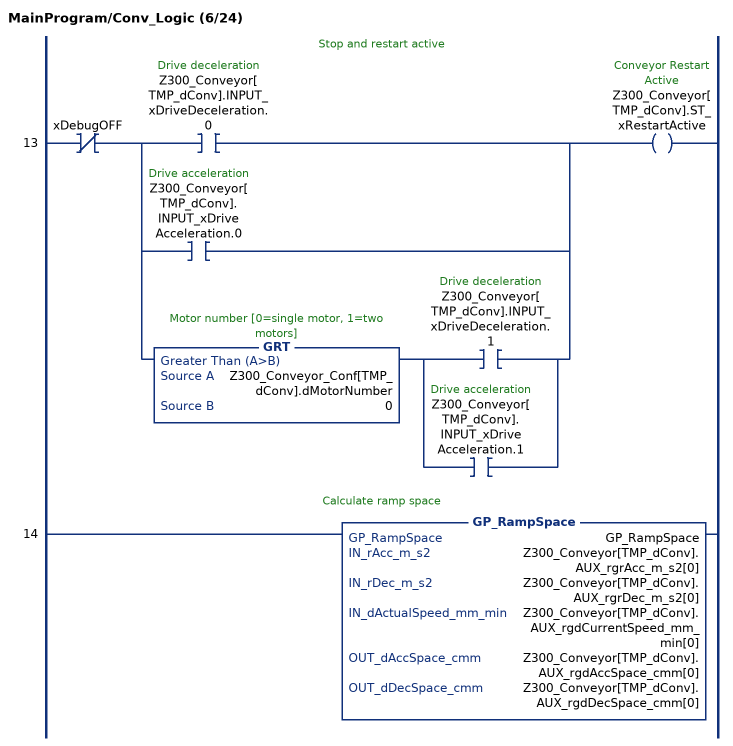
   // Stop and restart active
   13: XIO(xDebugOFF)[[XIC(Z300_Conveyor[TMP_dConv].INPUT_xDriveDeceleration.0) ,XIC(Z300_Conveyor[TMP_dConv].INPUT_xDriveAcceleration.0) ] ,GRT(Z300_Conveyor_Conf[TMP_dConv].dMotorNumber,0) [XIC(Z300_Conveyor[TMP_dConv].INPUT_xDriveDeceleration.1) ,XIC(Z300_Conveyor[TMP_dConv].INPUT_xDriveAcceleration.1) ] ]OTE(Z300_Conveyor[TMP_dConv].ST_xRestartActive);
   // Calculate ramp space
   14: GP_RampSpace(GP_RampSpace,Z300_Conveyor[TMP_dConv].AUX_rgrAcc_m_s2[0],Z300_Conveyor[TMP_dConv].AUX_rgrDec_m_s2[0],Z300_Conveyor[TMP_dConv].AUX_rgdCurrentSpeed_mm_min[0],Z300_Conveyor[TMP_dConv].AUX_rgdAccSpace_cmm[0],Z300_Conveyor[TMP_dConv].AUX_rgdDecSpace_cmm[0]);
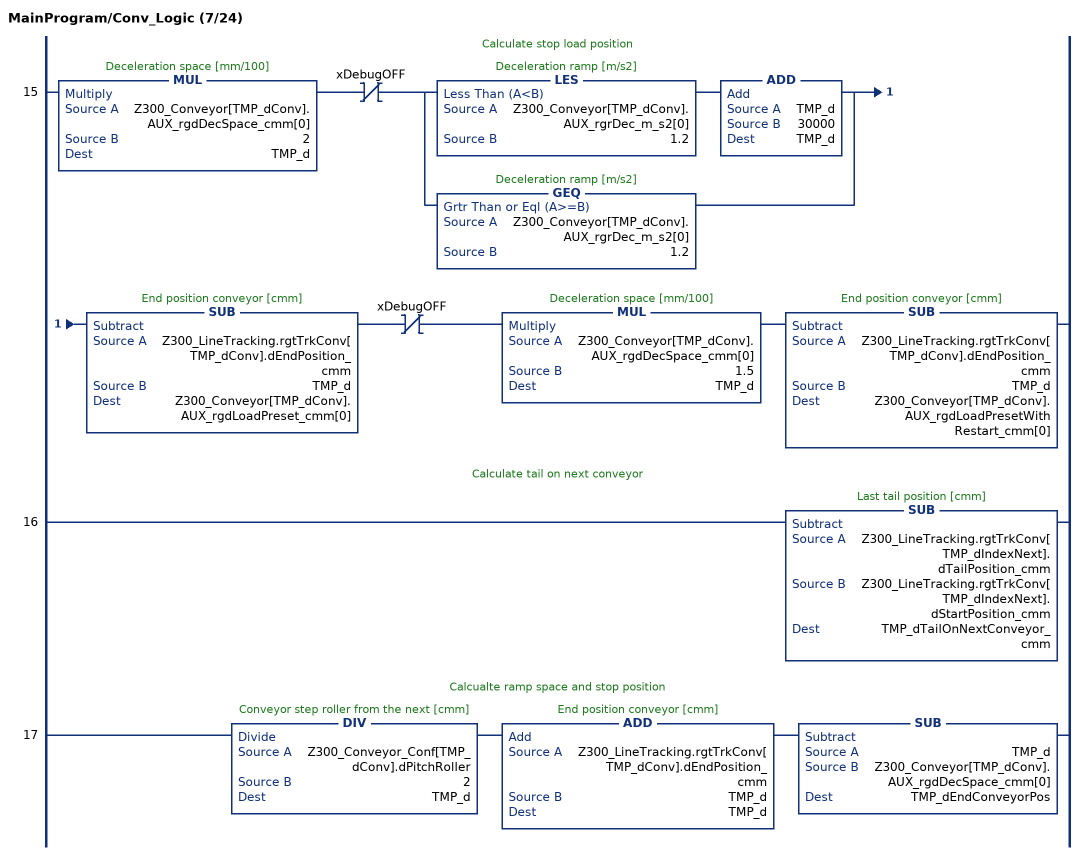
   // Calculate stop load position
   15: MUL(Z300_Conveyor[TMP_dConv].AUX_rgdDecSpace_cmm[0],2,TMP_d)XIO(xDebugOFF)[LES(Z300_Conveyor[TMP_dConv].AUX_rgrDec_m_s2[0],1.2) ADD(TMP_d,30000,TMP_d) ,GEQ(Z300_Conveyor[TMP_dConv].AUX_rgrDec_m_s2[0],1.2) ]SUB(Z300_LineTracking.rgtTrkConv[TMP_dConv].dEndPosition_cmm,TMP_d,Z300_Conveyor[TMP_dConv].AUX_rgdLoadPreset_cmm[0])XIO(xDebugOFF)MUL(Z300_Conveyor[TMP_dConv].AUX_rgdDecSpace_cmm[0],1.5,TMP_d)SUB(Z300_LineTracking.rgtTrkConv[TMP_dConv].dEndPosition_cmm,TMP_d,Z300_Conveyor[TMP_dConv].AUX_rgdLoadPresetWithRestart_cmm[0]);
   // Calculate tail on next conveyor
   16: SUB(Z300_LineTracking.rgtTrkConv[TMP_dIndexNext].dTailPosition_cmm,Z300_LineTracking.rgtTrkConv[TMP_dIndexNext].dStartPosition_cmm,TMP_dTailOnNextConveyor_cmm);
   // Calcualte ramp space and stop position
   17: DIV(Z300_Conveyor_Conf[TMP_dConv].dPitchRoller,2,TMP_d)ADD(Z300_LineTracking.rgtTrkConv[TMP_dConv].dEndPosition_cmm,TMP_d,TMP_d)SUB(TMP_d,Z300_Conveyor[TMP_dConv].AUX_rgdDecSpace_cmm[0],TMP_dEndConveyorPos);
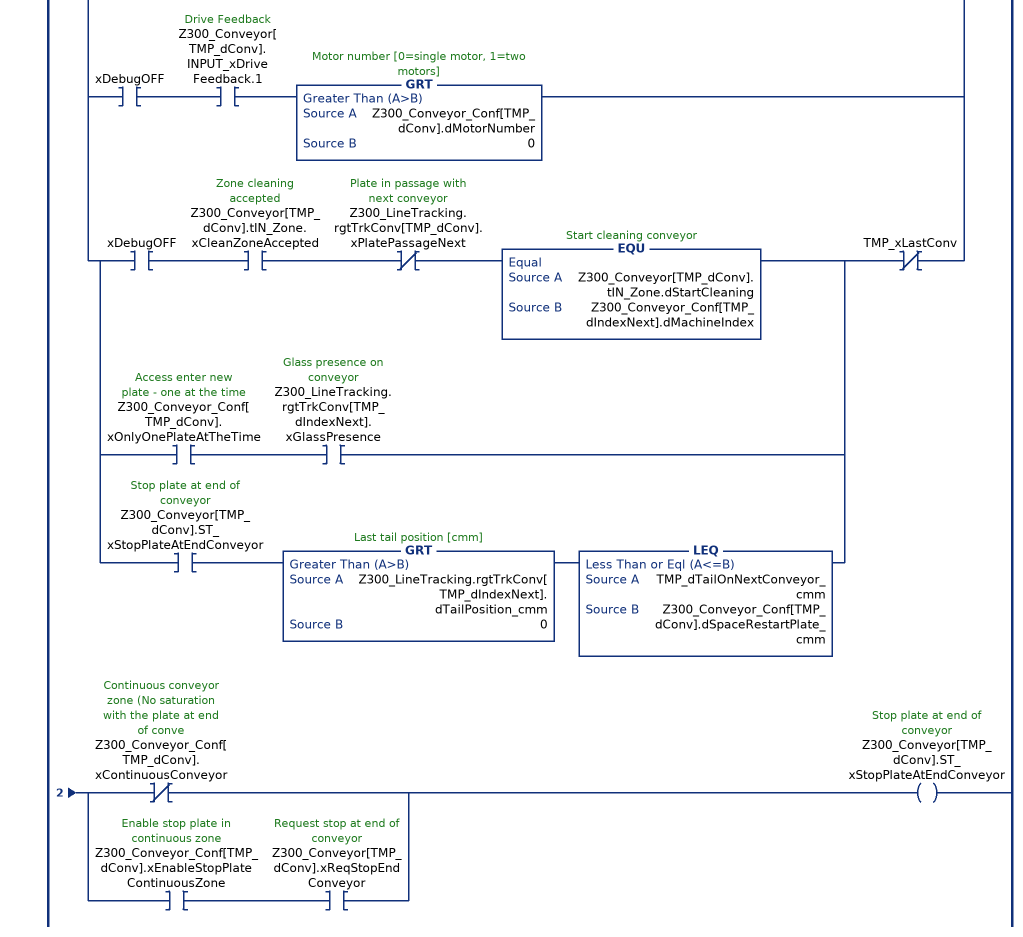
   // Stop at end of conveyor if next not run
   18: [GEQ(Z300_LineTracking.rgtTrkConv[TMP_dConv].dHeadPosition_cmm,Z300_Conveyor[TMP_dConv].AUX_rgdLoadPreset_cmm[0]) ,XIC(Z300_Conveyor[TMP_dConv].ST_xStopPlateAtEndConveyor) XIC(Z300_LineTracking.rgtTrkConv[TMP_dConv].xGlassPresCom) ][[XIO(Z300_Conveyor[TMP_dIndexNext].ST_xConveyorOutRun) ,XIC(xDebugON) ] [XIO(Z300_Conveyor[TMP_dIndexNext].ST_rgxConveyorOutRunSgm.0) ,XIO(Z300_Conveyor[TMP_dIndexNext].ST_rgxConveyorOutRunSgm.1) GRT(Z300_Conveyor_Conf[TMP_dIndexNext].dMotorNumber,0) ] XIO(TMP_xLastConv) ,XIC(Z300_Conveyor[TMP_dIndexNext].xReqExtStopLoadNewPlate) ,XIO(Z300_Conveyor[TMP_dConv].ST_xCleaningEnabled) XIC(Z300_Conveyor[TMP_dIndexNext].ST_xCleaningEnabled) XIO(Z300_LineTracking.rgtTrkConv[TMP_dConv].xPlatePassageNext) ,XIC(Z300_Conveyor[TMP_dConv].xReqStopEndConveyor) ,XIC(xDebugOFF) XIC(Z300_Conveyor[TMP_dConv].INPUT_xDriveFeedback.0) ,XIC(xDebugOFF) XIC(Z300_Conveyor[TMP_dConv].INPUT_xDriveFeedback.1) GRT(Z300_Conveyor_Conf[TMP_dConv].dMotorNumber,0) ,[XIC(xDebugOFF) XIC(Z300_Conveyor[TMP_dConv].tIN_Zone.xCleanZoneAccepted) XIO(Z300_LineTracking.rgtTrkConv[TMP_dConv].xPlatePassageNext) EQU(Z300_Conveyor[TMP_dConv].tIN_Zone.dStartCleaning,Z300_Conveyor_Conf[TMP_dIndexNext].dMachineIndex) ,XIC(Z300_Conveyor_Conf[TMP_dConv].xOnlyOnePlateAtTheTime) XIC(Z300_LineTracking.rgtTrkConv[TMP_dIndexNext].xGlassPresence) ,XIC(Z300_Conveyor[TMP_dConv].ST_xStopPlateAtEndConveyor) GRT(Z300_LineTracking.rgtTrkConv[TMP_dIndexNext].dTailPosition_cmm,0) LEQ(TMP_dTailOnNextConveyor_cmm,Z300_Conveyor_Conf[TMP_dConv].dSpaceRestartPlate_cmm) ] XIO(TMP_xLastConv) ][XIO(Z300_Conveyor_Conf[TMP_dConv].xContinuousConveyor) ,XIC(Z300_Conveyor_Conf[TMP_dConv].xEnableStopPlateContinuousZone) XIC(Z300_Conveyor[TMP_dConv].xReqStopEndConveyor) ]OTE(Z300_Conveyor[TMP_dConv].ST_xStopPlateAtEndConveyor);
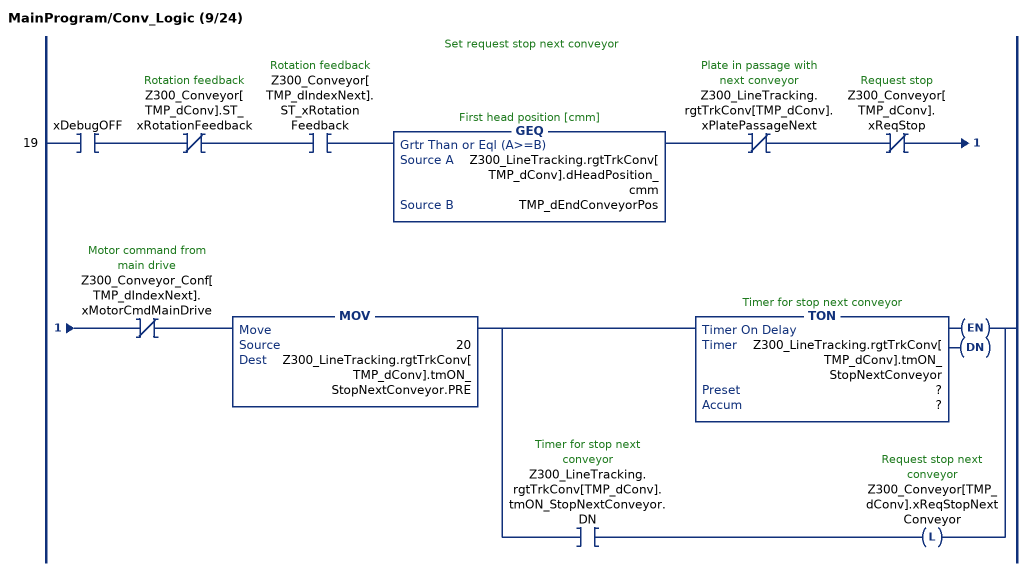
   // Set request stop next conveyor
   19: XIC(xDebugOFF)XIO(Z300_Conveyor[TMP_dConv].ST_xRotationFeedback)XIC(Z300_Conveyor[TMP_dIndexNext].ST_xRotationFeedback)GEQ(Z300_LineTracking.rgtTrkConv[TMP_dConv].dHeadPosition_cmm,TMP_dEndConveyorPos)XIO(Z300_LineTracking.rgtTrkConv[TMP_dConv].xPlatePassageNext)XIO(Z300_Conveyor[TMP_dConv].xReqStop)XIO(Z300_Conveyor_Conf[TMP_dIndexNext].xMotorCmdMainDrive)MOV(20,Z300_LineTracking.rgtTrkConv[TMP_dConv].tmON_StopNextConveyor.PRE)[TON(Z300_LineTracking.rgtTrkConv[TMP_dConv].tmON_StopNextConveyor,?,?) ,XIC(Z300_LineTracking.rgtTrkConv[TMP_dConv].tmON_StopNextConveyor.DN) OTL(Z300_Conveyor[TMP_dConv].xReqStopNextConveyor) ];
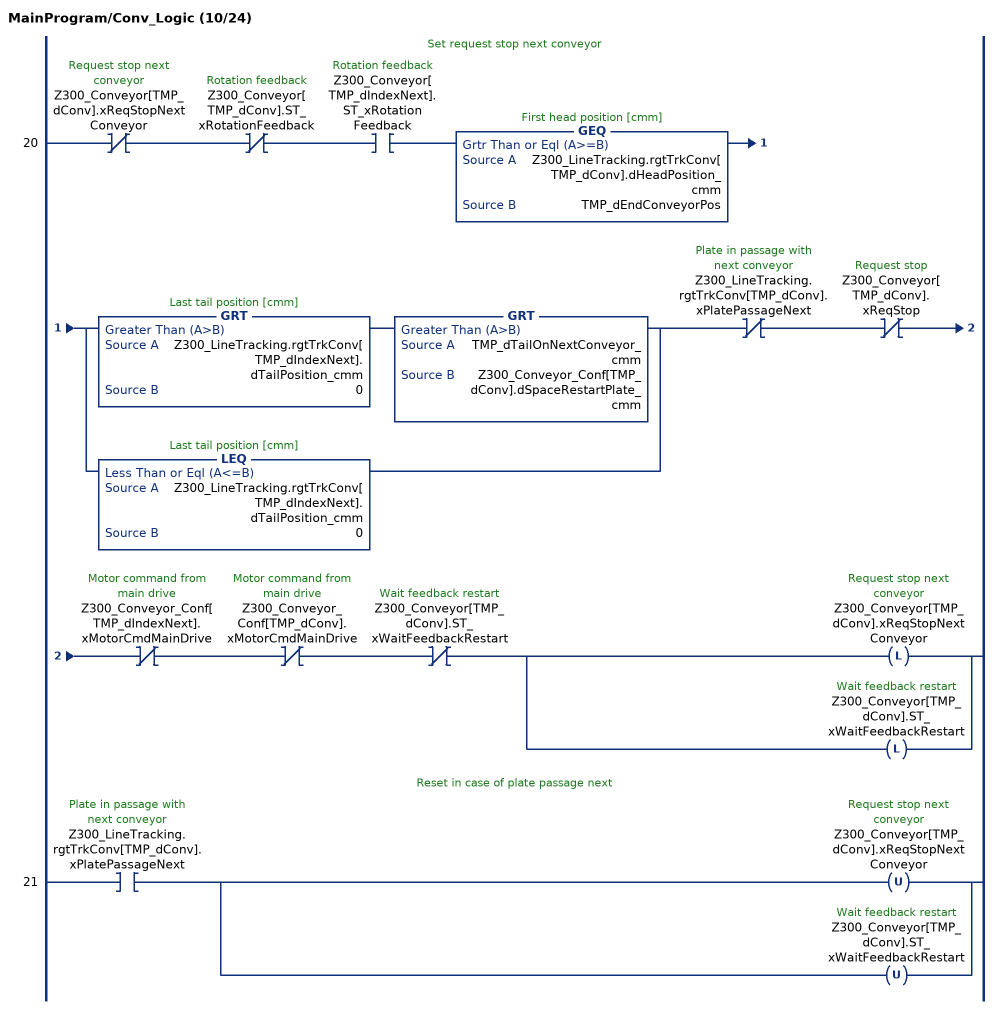
   // Set request stop next conveyor
   20: XIO(Z300_Conveyor[TMP_dConv].xReqStopNextConveyor)XIO(Z300_Conveyor[TMP_dConv].ST_xRotationFeedback)XIC(Z300_Conveyor[TMP_dIndexNext].ST_xRotationFeedback)GEQ(Z300_LineTracking.rgtTrkConv[TMP_dConv].dHeadPosition_cmm,TMP_dEndConveyorPos)[GRT(Z300_LineTracking.rgtTrkConv[TMP_dIndexNext].dTailPosition_cmm,0) GRT(TMP_dTailOnNextConveyor_cmm,Z300_Conveyor_Conf[TMP_dConv].dSpaceRestartPlate_cmm) ,LEQ(Z300_LineTracking.rgtTrkConv[TMP_dIndexNext].dTailPosition_cmm,0) ]XIO(Z300_LineTracking.rgtTrkConv[TMP_dConv].xPlatePassageNext)XIO(Z300_Conveyor[TMP_dConv].xReqStop)XIO(Z300_Conveyor_Conf[TMP_dIndexNext].xMotorCmdMainDrive)XIO(Z300_Conveyor_Conf[TMP_dConv].xMotorCmdMainDrive)XIO(Z300_Conveyor[TMP_dConv].ST_xWaitFeedbackRestart)[OTL(Z300_Conveyor[TMP_dConv].xReqStopNextConveyor) ,OTL(Z300_Conveyor[TMP_dConv].ST_xWaitFeedbackRestart) ];
   // Reset in case of plate passage next
   21: XIC(Z300_LineTracking.rgtTrkConv[TMP_dConv].xPlatePassageNext)[OTU(Z300_Conveyor[TMP_dConv].xReqStopNextConveyor) ,OTU(Z300_Conveyor[TMP_dConv].ST_xWaitFeedbackRestart) ];
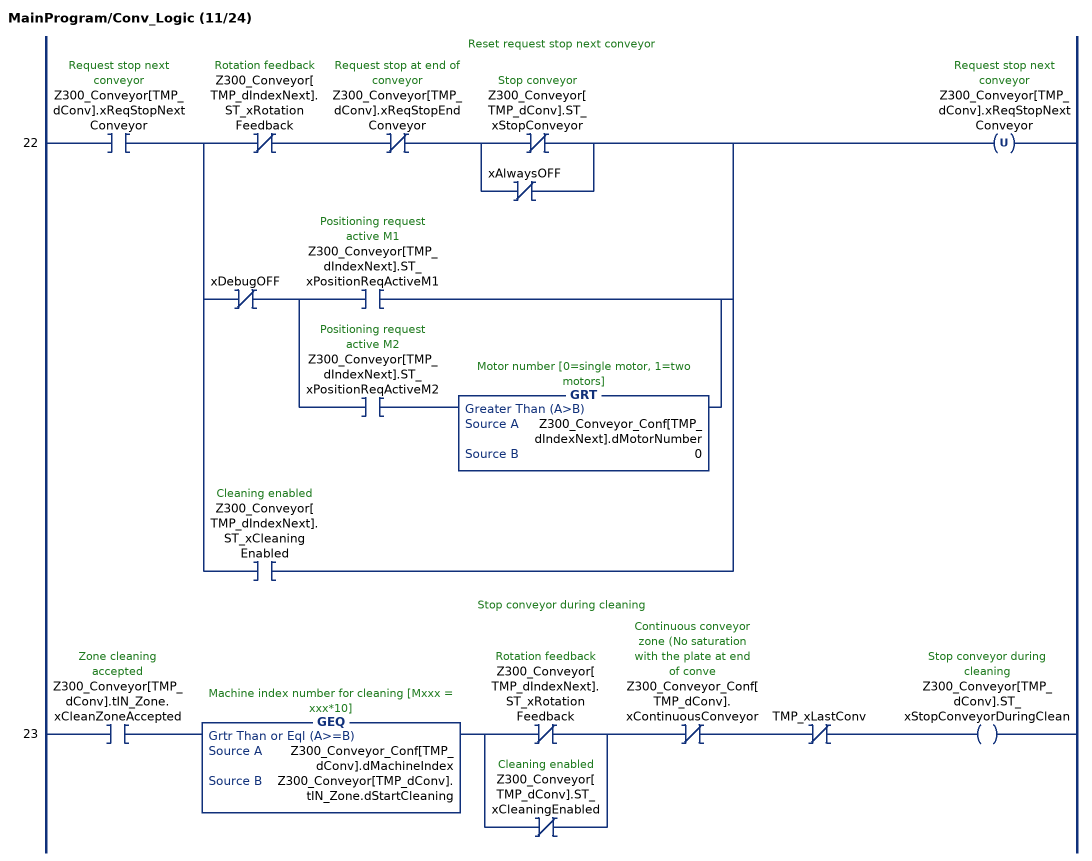
   // Reset request stop next conveyor
   22: XIC(Z300_Conveyor[TMP_dConv].xReqStopNextConveyor)[XIO(Z300_Conveyor[TMP_dIndexNext].ST_xRotationFeedback) XIO(Z300_Conveyor[TMP_dConv].xReqStopEndConveyor) [XIO(Z300_Conveyor[TMP_dConv].ST_xStopConveyor) ,XIO(xAlwaysOFF) ] ,XIO(xDebugOFF) [XIC(Z300_Conveyor[TMP_dIndexNext].ST_xPositionReqActiveM1) ,XIC(Z300_Conveyor[TMP_dIndexNext].ST_xPositionReqActiveM2) GRT(Z300_Conveyor_Conf[TMP_dIndexNext].dMotorNumber,0) ] ,XIC(Z300_Conveyor[TMP_dIndexNext].ST_xCleaningEnabled) ]OTU(Z300_Conveyor[TMP_dConv].xReqStopNextConveyor);
   // Stop conveyor during cleaning
   23: XIC(Z300_Conveyor[TMP_dConv].tIN_Zone.xCleanZoneAccepted)GEQ(Z300_Conveyor_Conf[TMP_dConv].dMachineIndex,Z300_Conveyor[TMP_dConv].tIN_Zone.dStartCleaning)[XIO(Z300_Conveyor[TMP_dIndexNext].ST_xRotationFeedback) ,XIO(Z300_Conveyor[TMP_dConv].ST_xCleaningEnabled) ]XIO(Z300_Conveyor_Conf[TMP_dConv].xContinuousConveyor)XIO(TMP_xLastConv)OTE(Z300_Conveyor[TMP_dConv].ST_xStopConveyorDuringClean);
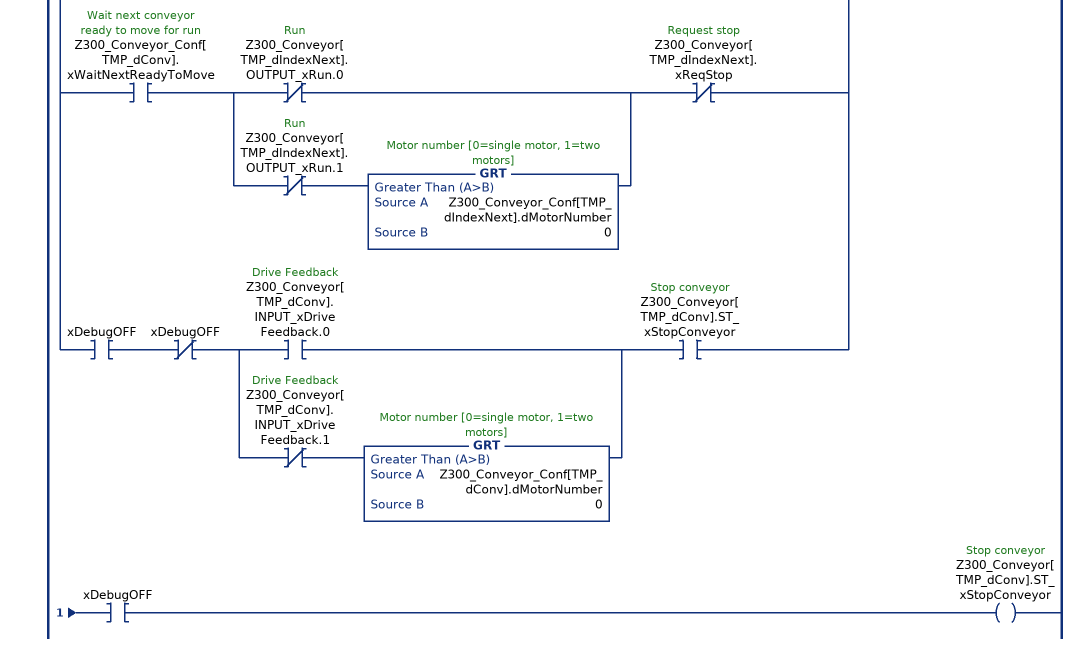
   // Stop conveyor
   24: [[XIC(Z300_LineTracking.rgtTrkConv[TMP_dConv].xPlatePassagePrevious) [XIO(Z300_Conveyor[TMP_dIndexPrevious].ST_xOutputEnable) ,XIC(Z300_Conveyor[TMP_dIndexPrevious].ST_xWaitStopConveyor) ,XIC(xAlwaysOFF) XIC(Z300_Conveyor[TMP_dIndexPrevious].xReqStop) ] ,XIC(Z300_LineTracking.rgtTrkConv[TMP_dConv].xPlatePassageNext) XIO(TMP_xLastConv) [XIO(Z300_Conveyor[TMP_dIndexNext].ST_xOutMotorRun) ,XIO(Z300_Conveyor[TMP_dIndexNext].INPUT_xSafetyConveyor) ] ,XIC(Z300_Conveyor[TMP_dConv].ST_xStopPlateAtEndConveyor) ,XIC(Z300_Conveyor[TMP_dConv].xReqStopNextConveyor) XIC(Z300_Conveyor[TMP_dIndexNext].ST_xRotationFeedback) ,XIC(Z300_Conveyor[TMP_dConv].ST_xStopConveyorDuringClean) ] [XIO(Z300_Conveyor_Conf[TMP_dConv].xContinuousConveyor) ,XIC(Z300_Conveyor_Conf[TMP_dConv].xEnableStopPlateContinuousZone) XIC(Z300_Conveyor[TMP_dConv].xReqStopEndConveyor) ] ,XIC(Z300_Conveyor[TMP_dIndexPrevious].xReqStopNextConveyor) XIO(Z300_Conveyor[TMP_dConv].tIN_Zone.xCleanZoneAccepted) XIO(Z300_LineTracking.rgtTrkConv[TMP_dConv].xGlassPresence) ,XIC(Z300_Conveyor_Conf[TMP_dConv].xWaitNextReadyToMove) [XIO(Z300_Conveyor[TMP_dIndexNext].OUTPUT_xRun.0) ,XIO(Z300_Conveyor[TMP_dIndexNext].OUTPUT_xRun.1) GRT(Z300_Conveyor_Conf[TMP_dIndexNext].dMotorNumber,0) ] XIO(Z300_Conveyor[TMP_dIndexNext].xReqStop) ,XIC(xDebugOFF) XIO(xDebugOFF) [XIC(Z300_Conveyor[TMP_dConv].INPUT_xDriveFeedback.0) ,XIO(Z300_Conveyor[TMP_dConv].INPUT_xDriveFeedback.1) GRT(Z300_Conveyor_Conf[TMP_dConv].dMotorNumber,0) ] XIC(Z300_Conveyor[TMP_dConv].ST_xStopConveyor) ]XIO(Z300_Conveyor[TMP_dConv].xReqBypassEndStop)XIC(xDebugOFF)OTE(Z300_Conveyor[TMP_dConv].ST_xStopConveyor);
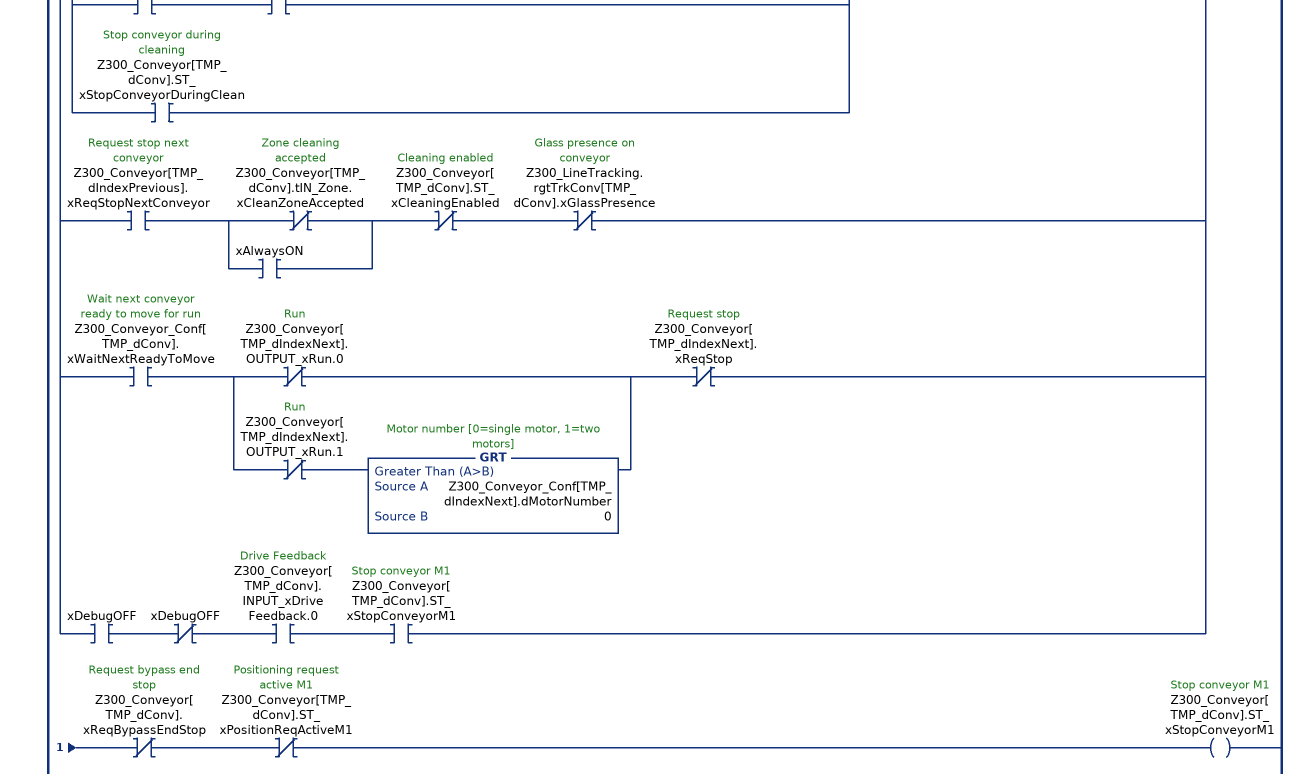
   // Stop conveyor M1
   // Monterrey VF2 - If this is conveyor after drop section I stop convveyor just if tail is under certain quote
   25: [[XIC(Z300_LineTracking.rgtTrkConv[TMP_dConv].xPlatePassagePrevious) [XIO(Z300_Conveyor[TMP_dIndexPrevious].ST_xOutputEnable) ,XIC(xDebugOFF) XIO(Z300_Conveyor[TMP_dIndexPrevious].tmON_DelayReadyToMove[0].DN) ,XIC(Z300_Conveyor[TMP_dIndexPrevious].ST_xInitialCondition) ,XIC(xDebugOFF) XIC(Z300_Conveyor[TMP_dIndexPrevious].ST_xWaitStopConveyor) ,XIC(xAlwaysOFF) XIC(Z300_Conveyor[TMP_dIndexPrevious].xReqStop) ] ,XIC(Z300_LineTracking.rgtTrkConv[TMP_dConv].xPlatePassageNext) XIO(TMP_xLastConv) [[XIO(Z300_Conveyor[TMP_dIndexNext].ST_xOutMotorRun) ,XIC(xAlwaysON) ] XIO(Z300_Conveyor[TMP_dIndexNext].ST_rgxConveyorOutRunSgm.0) XIO(Z300_Conveyor[TMP_dIndexNext].ST_rgxConveyorOutRunSgm.1) ,XIO(Z300_Conveyor[TMP_dIndexNext].INPUT_xSafetyConveyor) ] ,XIC(Z300_Conveyor[TMP_dConv].ST_xStopPlateAtEndConveyor) XIO(Z300_Conveyor[TMP_dConv].xReqBypassEndConveyorM1) ,XIC(Z300_Conveyor[TMP_dConv].xReqStopNextConveyor) XIC(Z300_Conveyor[TMP_dIndexNext].ST_xRotationFeedback) ,XIC(Z300_Conveyor[TMP_dConv].ST_xStopConveyorDuringClean) ] [XIO(Z300_Conveyor_Conf[TMP_dConv].xContinuousConveyor) ,XIC(Z300_Conveyor_Conf[TMP_dConv].xEnableStopPlateContinuousZone) XIC(Z300_Conveyor[TMP_dConv].xReqStopEndConveyor) ] ,XIC(Z300_Conveyor[TMP_dIndexPrevious].xReqStopNextConveyor) [XIO(Z300_Conveyor[TMP_dConv].tIN_Zone.xCleanZoneAccepted) ,XIC(xAlwaysON) ] XIO(Z300_Conveyor[TMP_dConv].ST_xCleaningEnabled) XIO(Z300_LineTracking.rgtTrkConv[TMP_dConv].xGlassPresence) ,XIC(Z300_Conveyor_Conf[TMP_dConv].xWaitNextReadyToMove) [XIO(Z300_Conveyor[TMP_dIndexNext].OUTPUT_xRun.0) ,XIO(Z300_Conveyor[TMP_dIndexNext].OUTPUT_xRun.1) GRT(Z300_Conveyor_Conf[TMP_dIndexNext].dMotorNumber,0) ] XIO(Z300_Conveyor[TMP_dIndexNext].xReqStop) ,XIC(xDebugOFF) XIO(xDebugOFF) XIC(Z300_Conveyor[TMP_dConv].INPUT_xDriveFeedback.0) XIC(Z300_Conveyor[TMP_dConv].ST_xStopConveyorM1) ]XIO(Z300_Conveyor[TMP_dConv].xReqBypassEndStop)XIO(Z300_Conveyor[TMP_dConv].ST_xPositionReqActiveM1)OTE(Z300_Conveyor[TMP_dConv].ST_xStopConveyorM1);
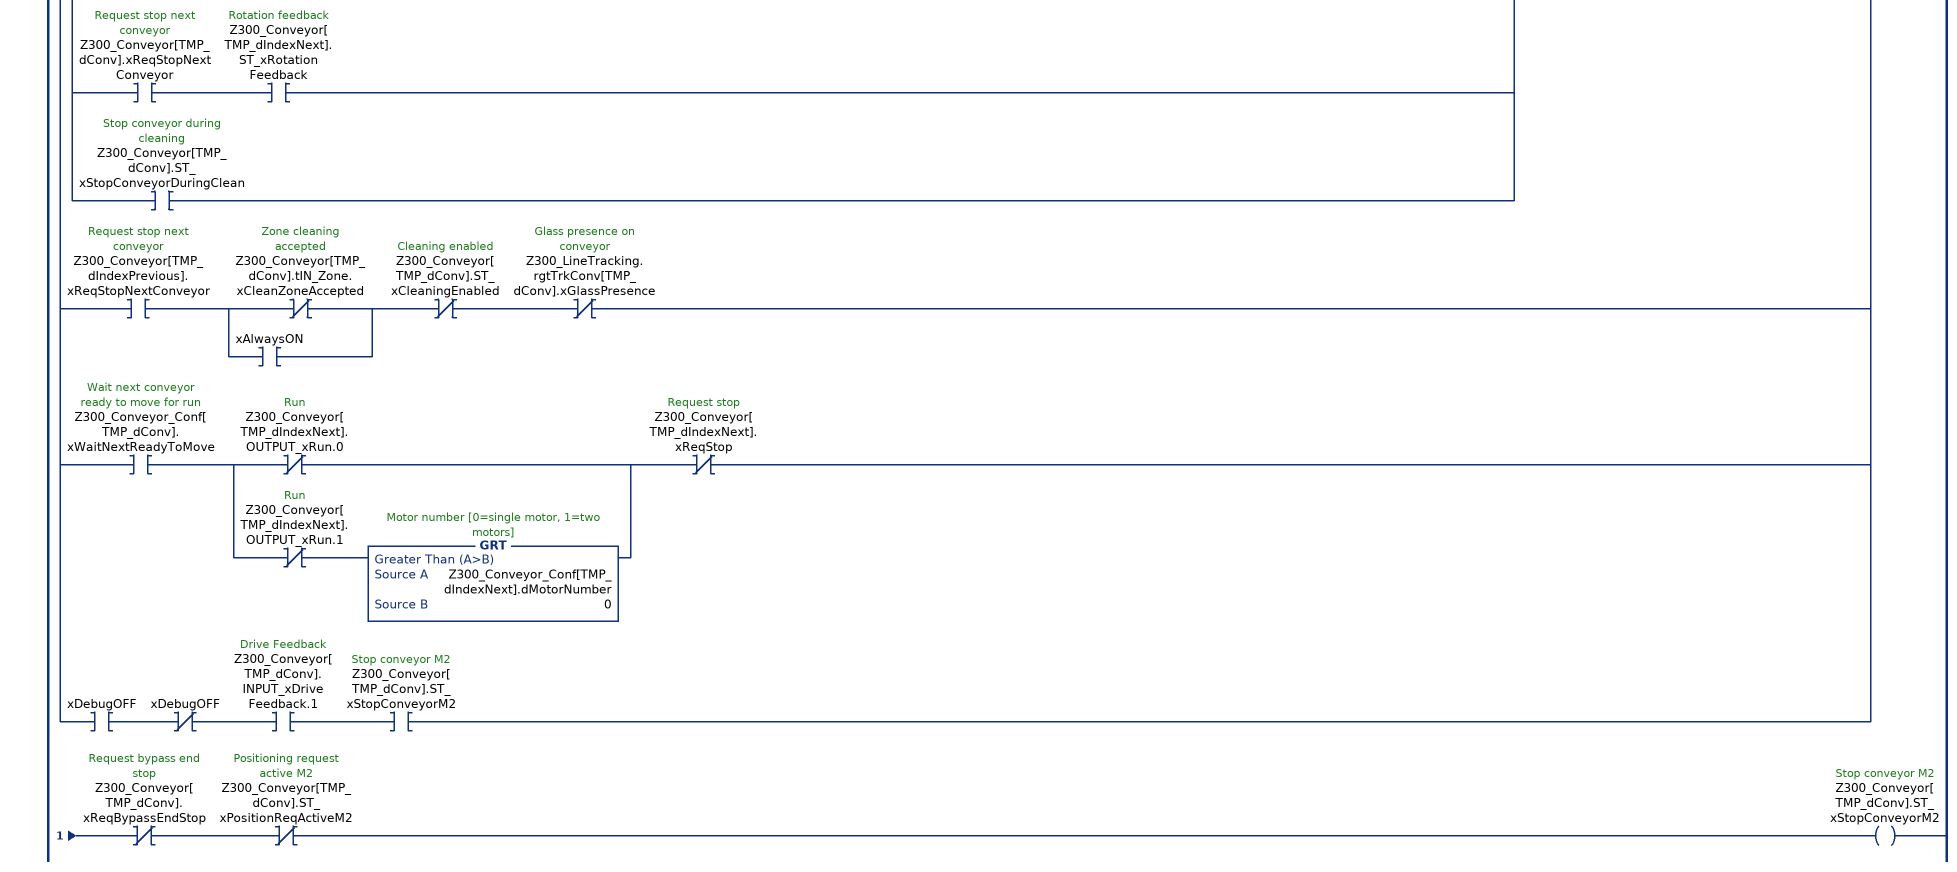
   // Stop conveyor M2
   // Monterrey VF2 - If this is conveyor after drop section I stop convveyor just if tail is under certain quote
   26: [[XIC(Z300_LineTracking.rgtTrkConv[TMP_dConv].xPlatePassagePrevious) [XIO(Z300_Conveyor[TMP_dIndexPrevious].ST_xOutputEnable) ,XIC(xDebugOFF) XIO(Z300_Conveyor[TMP_dIndexPrevious].tmON_DelayReadyToMove[1].DN) ,XIC(Z300_Conveyor[TMP_dIndexPrevious].ST_xInitialCondition) ,XIC(xDebugOFF) XIC(Z300_Conveyor[TMP_dIndexPrevious].ST_xWaitStopConveyor) ,XIC(xAlwaysOFF) XIC(Z300_Conveyor[TMP_dIndexPrevious].xReqStop) ] ,XIC(Z300_LineTracking.rgtTrkConv[TMP_dConv].xPlatePassageNext) XIO(TMP_xLastConv) [XIO(xDebugOFF) [EQU(TMP_dConv,12) LES(Z300_LineTracking.rgtTrkConv[TMP_dConv].dTailPosition_cmm,4100000) ,NEQ(TMP_dConv,12) ] XIO(xDebugOFF) [XIO(Z300_Conveyor[TMP_dIndexNext].ST_xOutMotorRun) ,XIC(xAlwaysON) ] XIO(Z300_Conveyor[TMP_dIndexNext].ST_rgxConveyorOutRunSgm.0) XIO(Z300_Conveyor[TMP_dIndexNext].ST_rgxConveyorOutRunSgm.1) ,XIO(Z300_Conveyor[TMP_dIndexNext].INPUT_xSafetyConveyor) ] ,XIC(Z300_Conveyor[TMP_dConv].ST_xStopPlateAtEndConveyor) XIO(Z300_Conveyor[TMP_dConv].xReqBypassEndConveyorM2) ,XIC(Z300_Conveyor[TMP_dConv].xReqStopNextConveyor) XIC(Z300_Conveyor[TMP_dIndexNext].ST_xRotationFeedback) ,XIC(Z300_Conveyor[TMP_dConv].ST_xStopConveyorDuringClean) ] [XIO(Z300_Conveyor_Conf[TMP_dConv].xContinuousConveyor) ,XIC(Z300_Conveyor_Conf[TMP_dConv].xEnableStopPlateContinuousZone) XIC(Z300_Conveyor[TMP_dConv].xReqStopEndConveyor) ] ,XIC(Z300_Conveyor[TMP_dIndexPrevious].xReqStopNextConveyor) [XIO(Z300_Conveyor[TMP_dConv].tIN_Zone.xCleanZoneAccepted) ,XIC(xAlwaysON) ] XIO(Z300_Conveyor[TMP_dConv].ST_xCleaningEnabled) XIO(Z300_LineTracking.rgtTrkConv[TMP_dConv].xGlassPresence) ,XIC(Z300_Conveyor_Conf[TMP_dConv].xWaitNextReadyToMove) [XIO(Z300_Conveyor[TMP_dIndexNext].OUTPUT_xRun.0) ,XIO(Z300_Conveyor[TMP_dIndexNext].OUTPUT_xRun.1) GRT(Z300_Conveyor_Conf[TMP_dIndexNext].dMotorNumber,0) ] XIO(Z300_Conveyor[TMP_dIndexNext].xReqStop) ,XIC(xDebugOFF) XIO(xDebugOFF) XIC(Z300_Conveyor[TMP_dConv].INPUT_xDriveFeedback.1) XIC(Z300_Conveyor[TMP_dConv].ST_xStopConveyorM2) ]XIO(Z300_Conveyor[TMP_dConv].xReqBypassEndStop)XIO(Z300_Conveyor[TMP_dConv].ST_xPositionReqActiveM2)OTE(Z300_Conveyor[TMP_dConv].ST_xStopConveyorM2);
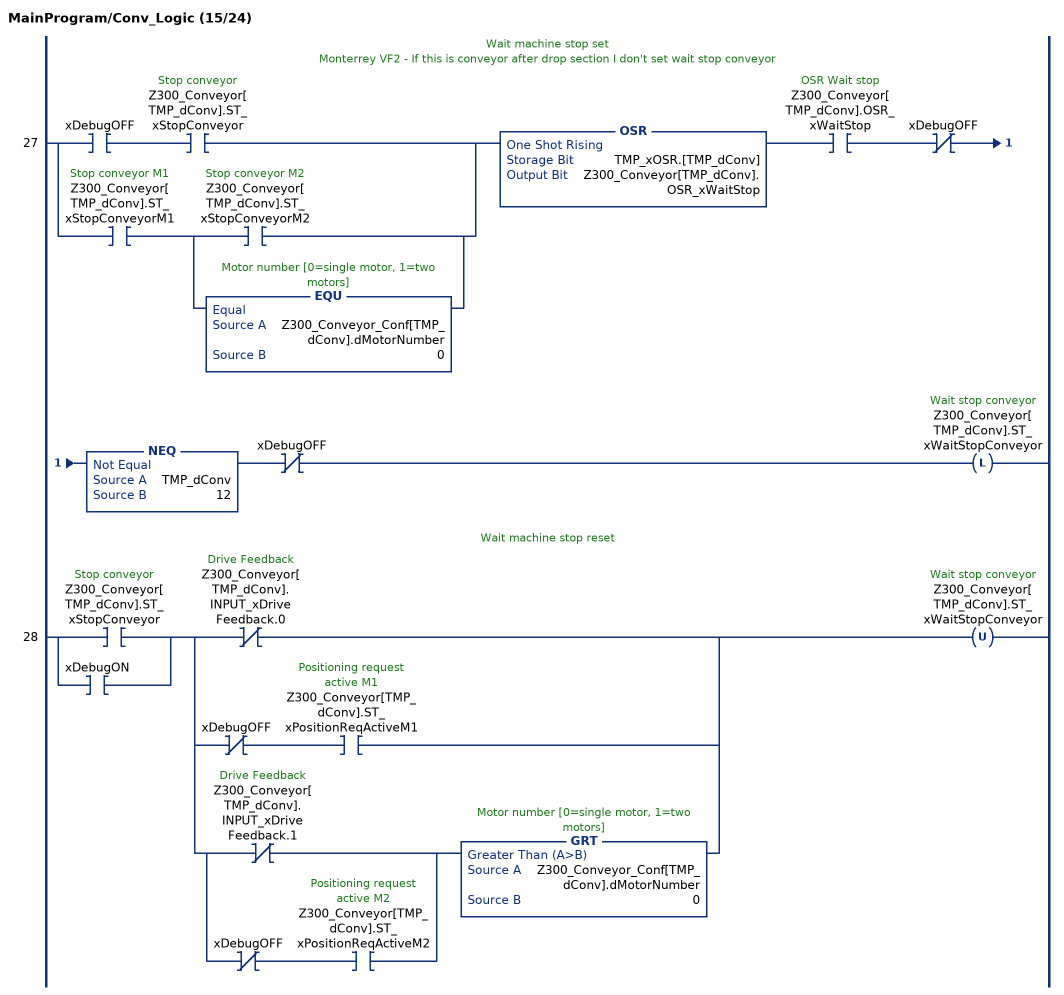
   // Wait machine stop set
   // Monterrey VF2 - If this is conveyor after drop section I don't set wait stop conveyor
   27: [XIC(xDebugOFF) XIC(Z300_Conveyor[TMP_dConv].ST_xStopConveyor) ,XIC(Z300_Conveyor[TMP_dConv].ST_xStopConveyorM1) [XIC(Z300_Conveyor[TMP_dConv].ST_xStopConveyorM2) ,EQU(Z300_Conveyor_Conf[TMP_dConv].dMotorNumber,0) ] ]OSR(TMP_xOSR.[TMP_dConv],Z300_Conveyor[TMP_dConv].OSR_xWaitStop)XIC(Z300_Conveyor[TMP_dConv].OSR_xWaitStop)XIO(xDebugOFF)NEQ(TMP_dConv,12)XIO(xDebugOFF)OTL(Z300_Conveyor[TMP_dConv].ST_xWaitStopConveyor);
   // Wait machine stop reset
   28: [XIC(Z300_Conveyor[TMP_dConv].ST_xStopConveyor) ,XIC(xDebugON) ][[XIO(Z300_Conveyor[TMP_dConv].INPUT_xDriveFeedback.0) ,XIO(xDebugOFF) XIC(Z300_Conveyor[TMP_dConv].ST_xPositionReqActiveM1) ] ,[XIO(Z300_Conveyor[TMP_dConv].INPUT_xDriveFeedback.1) ,XIO(xDebugOFF) XIC(Z300_Conveyor[TMP_dConv].ST_xPositionReqActiveM2) ] GRT(Z300_Conveyor_Conf[TMP_dConv].dMotorNumber,0) ]OTU(Z300_Conveyor[TMP_dConv].ST_xWaitStopConveyor);
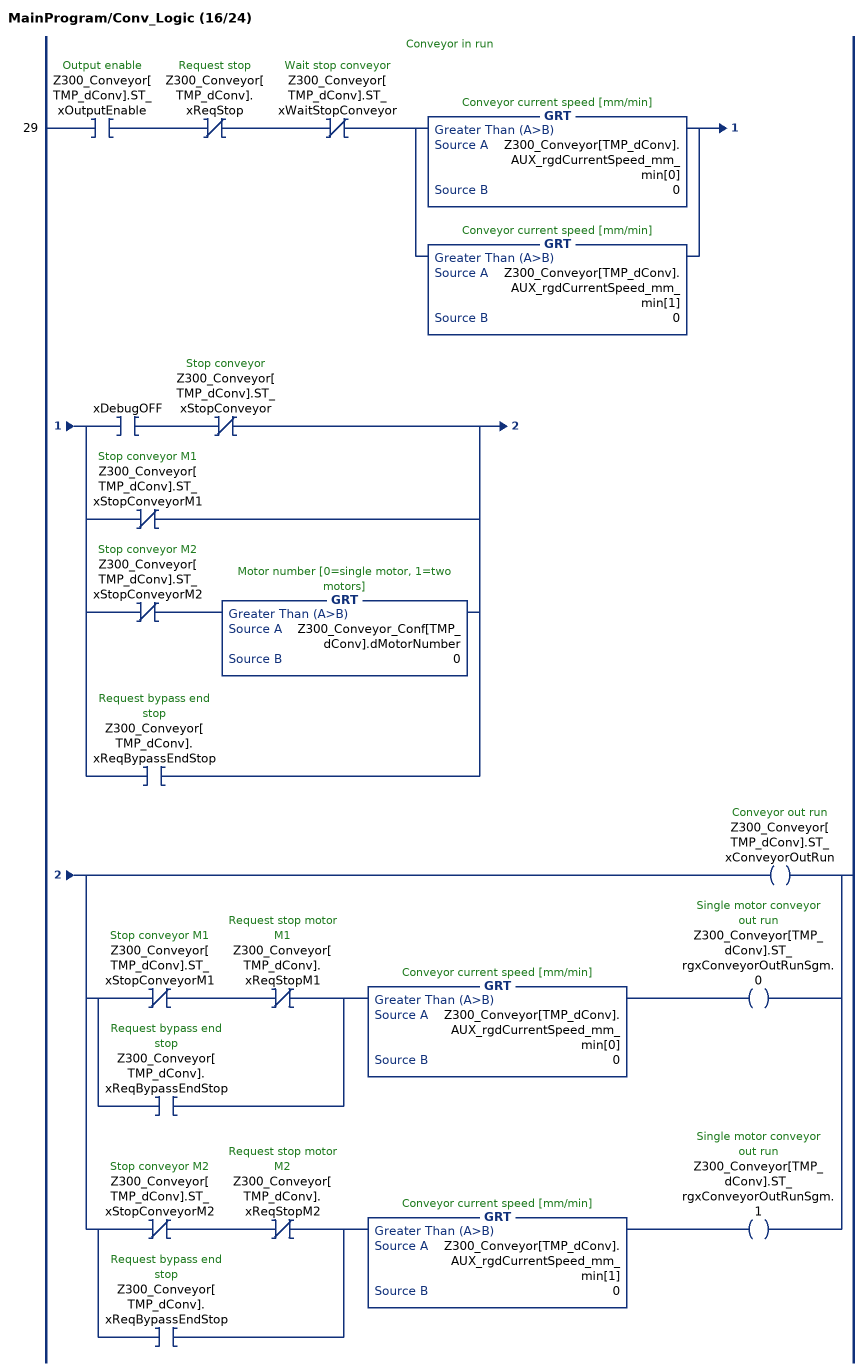
   // Conveyor in run
   29: XIC(Z300_Conveyor[TMP_dConv].ST_xOutputEnable)XIO(Z300_Conveyor[TMP_dConv].xReqStop)XIO(Z300_Conveyor[TMP_dConv].ST_xWaitStopConveyor)[GRT(Z300_Conveyor[TMP_dConv].AUX_rgdCurrentSpeed_mm_min[0],0) ,GRT(Z300_Conveyor[TMP_dConv].AUX_rgdCurrentSpeed_mm_min[1],0) ][XIC(xDebugOFF) XIO(Z300_Conveyor[TMP_dConv].ST_xStopConveyor) ,XIO(Z300_Conveyor[TMP_dConv].ST_xStopConveyorM1) ,XIO(Z300_Conveyor[TMP_dConv].ST_xStopConveyorM2) GRT(Z300_Conveyor_Conf[TMP_dConv].dMotorNumber,0) ,XIC(Z300_Conveyor[TMP_dConv].xReqBypassEndStop) ][OTE(Z300_Conveyor[TMP_dConv].ST_xConveyorOutRun) ,[XIO(Z300_Conveyor[TMP_dConv].ST_xStopConveyorM1) XIO(Z300_Conveyor[TMP_dConv].xReqStopM1) ,XIC(Z300_Conveyor[TMP_dConv].xReqBypassEndStop) ] GRT(Z300_Conveyor[TMP_dConv].AUX_rgdCurrentSpeed_mm_min[0],0) OTE(Z300_Conveyor[TMP_dConv].ST_rgxConveyorOutRunSgm.0) ,[XIO(Z300_Conveyor[TMP_dConv].ST_xStopConveyorM2) XIO(Z300_Conveyor[TMP_dConv].xReqStopM2) ,XIC(Z300_Conveyor[TMP_dConv].xReqBypassEndStop) ] GRT(Z300_Conveyor[TMP_dConv].AUX_rgdCurrentSpeed_mm_min[1],0) OTE(Z300_Conveyor[TMP_dConv].ST_rgxConveyorOutRunSgm.1) ];
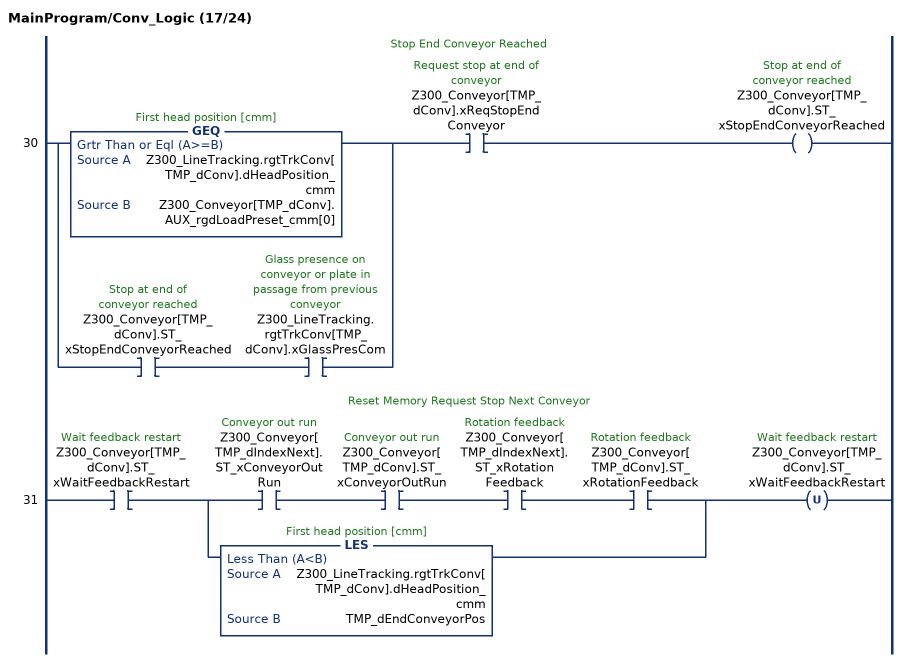
   // Stop End Conveyor Reached
   30: [GEQ(Z300_LineTracking.rgtTrkConv[TMP_dConv].dHeadPosition_cmm,Z300_Conveyor[TMP_dConv].AUX_rgdLoadPreset_cmm[0]) ,XIC(Z300_Conveyor[TMP_dConv].ST_xStopEndConveyorReached) XIC(Z300_LineTracking.rgtTrkConv[TMP_dConv].xGlassPresCom) ]XIC(Z300_Conveyor[TMP_dConv].xReqStopEndConveyor)OTE(Z300_Conveyor[TMP_dConv].ST_xStopEndConveyorReached);
   // Reset Memory Request Stop Next Conveyor
   31: XIC(Z300_Conveyor[TMP_dConv].ST_xWaitFeedbackRestart)[XIC(Z300_Conveyor[TMP_dIndexNext].ST_xConveyorOutRun) XIC(Z300_Conveyor[TMP_dConv].ST_xConveyorOutRun) XIC(Z300_Conveyor[TMP_dIndexNext].ST_xRotationFeedback) XIC(Z300_Conveyor[TMP_dConv].ST_xRotationFeedback) ,LES(Z300_LineTracking.rgtTrkConv[TMP_dConv].dHeadPosition_cmm,TMP_dEndConveyorPos) ]OTU(Z300_Conveyor[TMP_dConv].ST_xWaitFeedbackRestart);
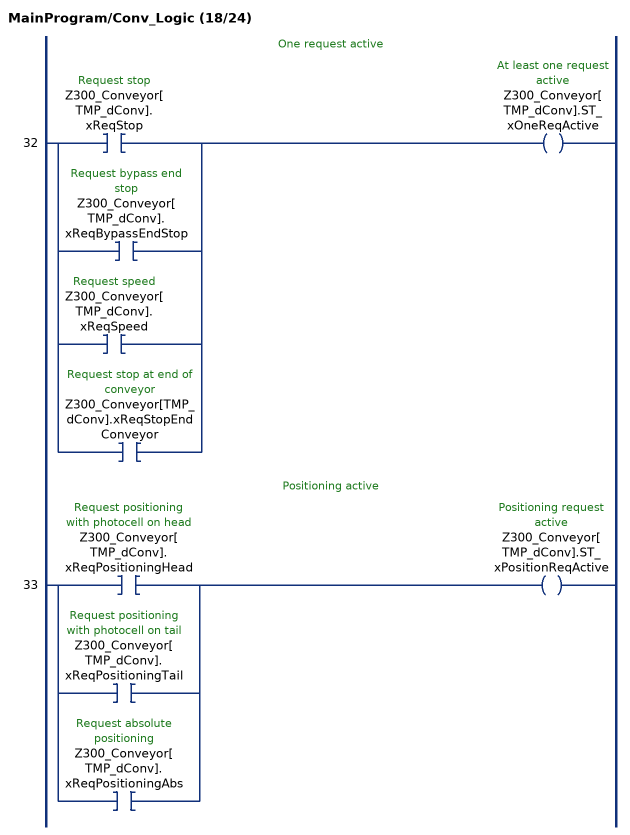
   // One request active
   32: [XIC(Z300_Conveyor[TMP_dConv].xReqStop) ,XIC(Z300_Conveyor[TMP_dConv].xReqBypassEndStop) ,XIC(Z300_Conveyor[TMP_dConv].xReqSpeed) ,XIC(Z300_Conveyor[TMP_dConv].xReqStopEndConveyor) ]OTE(Z300_Conveyor[TMP_dConv].ST_xOneReqActive);
   // Positioning active
   33: [XIC(Z300_Conveyor[TMP_dConv].xReqPositioningHead) ,XIC(Z300_Conveyor[TMP_dConv].xReqPositioningTail) ,XIC(Z300_Conveyor[TMP_dConv].xReqPositioningAbs) ]OTE(Z300_Conveyor[TMP_dConv].ST_xPositionReqActive);
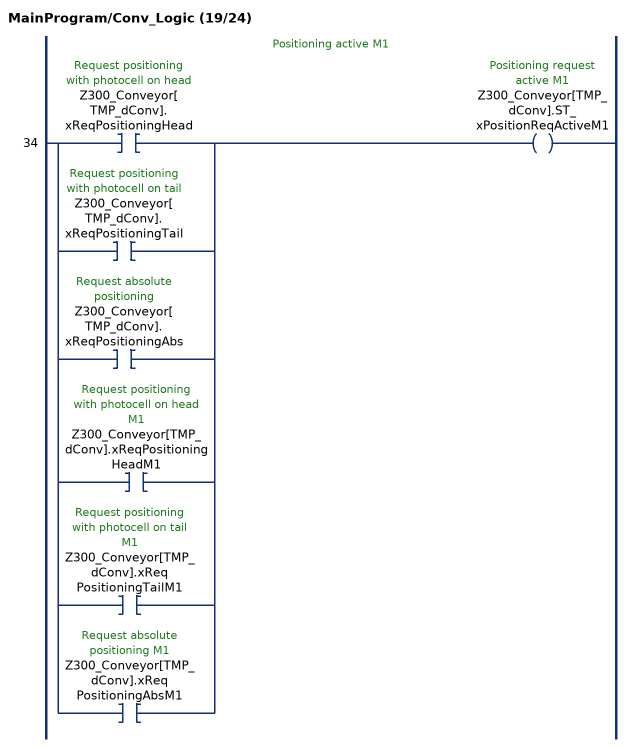
   // Positioning active M1
   34: [XIC(Z300_Conveyor[TMP_dConv].xReqPositioningHead) ,XIC(Z300_Conveyor[TMP_dConv].xReqPositioningTail) ,XIC(Z300_Conveyor[TMP_dConv].xReqPositioningAbs) ,XIC(Z300_Conveyor[TMP_dConv].xReqPositioningHeadM1) ,XIC(Z300_Conveyor[TMP_dConv].xReqPositioningTailM1) ,XIC(Z300_Conveyor[TMP_dConv].xReqPositioningAbsM1) ]OTE(Z300_Conveyor[TMP_dConv].ST_xPositionReqActiveM1);
